REGION Network 268
   RUNG wire#powerrail
      Contact( "EMS".Carrier[02].SDC_OUT.HeartBeat )
      Coil( "Carrier_02_Heartbeat" )
   END_RUNG
   // the same network as SCL:
   "Carrier_02_Heartbeat" := "EMS".Carrier[02].SDC_OUT.HeartBeat;
END_REGION

REGION Network 269
   RUNG wire#powerrail
      Contact( "EMS".Carrier[02].SDC_OUT.DriveFwdCMD )
      I_Contact( "EMS".Carrier[01].SDC_IN.CrashDetectStatus )
      Coil( "Carrier_02_Drive_Forward_Command" )
   END_RUNG
   // the same network as SCL:
   "Carrier_02_Drive_Forward_Command" := "EMS".Carrier[02].SDC_OUT.DriveFwdCMD AND NOT "EMS".Carrier[01].SDC_IN.CrashDetectStatus;
END_REGION

REGION Network 270
   RUNG wire#powerrail
      Contact( "EMS".Carrier[02].SDC_OUT.FaultReset )
      Coil( "Carrier_02_Fault_Reset" )
   END_RUNG
   // the same network as SCL:
   "Carrier_02_Fault_Reset" := "EMS".Carrier[02].SDC_OUT.FaultReset;
END_REGION

REGION Network 271
   RUNG wire#powerrail
      Contact( "EMS".Carrier[02].SDC_OUT.AtCmdPos )
      Coil( "Carrier_02_At_Command_Position" )
   END_RUNG
   // the same network as SCL:
   "Carrier_02_At_Command_Position" := "EMS".Carrier[02].SDC_OUT.AtCmdPos;
END_REGION

REGION Network 272
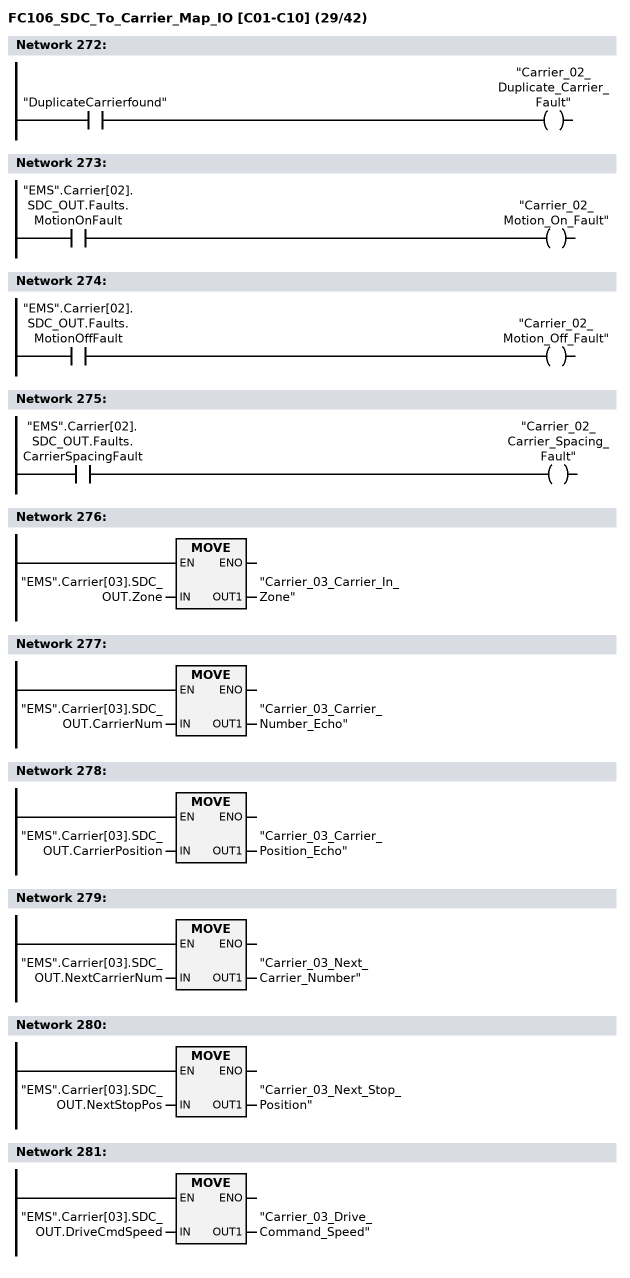
   RUNG wire#powerrail
      Contact( "DuplicateCarrierfound" )
      Coil( "Carrier_02_Duplicate_Carrier_Fault" )
   END_RUNG
   // the same network as SCL:
   "Carrier_02_Duplicate_Carrier_Fault" := "DuplicateCarrierfound";
END_REGION

REGION Network 273
   RUNG wire#powerrail
      Contact( "EMS".Carrier[02].SDC_OUT.Faults.MotionOnFault )
      Coil( "Carrier_02_Motion_On_Fault" )
   END_RUNG
   // the same network as SCL:
   "Carrier_02_Motion_On_Fault" := "EMS".Carrier[02].SDC_OUT.Faults.MotionOnFault;
END_REGION

REGION Network 274
   RUNG wire#powerrail
      Contact( "EMS".Carrier[02].SDC_OUT.Faults.MotionOffFault )
      Coil( "Carrier_02_Motion_Off_Fault" )
   END_RUNG
   // the same network as SCL:
   "Carrier_02_Motion_Off_Fault" := "EMS".Carrier[02].SDC_OUT.Faults.MotionOffFault;
END_REGION

REGION Network 275
   RUNG wire#powerrail
      Contact( "EMS".Carrier[02].SDC_OUT.Faults.CarrierSpacingFault )
      Coil( "Carrier_02_Carrier_Spacing_Fault" )
   END_RUNG
   // the same network as SCL:
   "Carrier_02_Carrier_Spacing_Fault" := "EMS".Carrier[02].SDC_OUT.Faults.CarrierSpacingFault;
END_REGION

REGION Network 276
   RUNG wire#powerrail
      Move(in := "EMS".Carrier[03].SDC_OUT.Zone, out1 => "Carrier_03_Carrier_In_Zone")
   END_RUNG
   // the same network as SCL:
   "Carrier_03_Carrier_In_Zone" := "EMS".Carrier[03].SDC_OUT.Zone;
END_REGION

REGION Network 277
   RUNG wire#powerrail
      Move(in := "EMS".Carrier[03].SDC_OUT.CarrierNum, out1 => "Carrier_03_Carrier_Number_Echo")
   END_RUNG
   // the same network as SCL:
   "Carrier_03_Carrier_Number_Echo" := "EMS".Carrier[03].SDC_OUT.CarrierNum;
END_REGION

REGION Network 278
   RUNG wire#powerrail
      Move(in := "EMS".Carrier[03].SDC_OUT.CarrierPosition, out1 => "Carrier_03_Carrier_Position_Echo")
   END_RUNG
   // the same network as SCL:
   "Carrier_03_Carrier_Position_Echo" := "EMS".Carrier[03].SDC_OUT.CarrierPosition;
END_REGION

REGION Network 279
   RUNG wire#powerrail
      Move(in := "EMS".Carrier[03].SDC_OUT.NextCarrierNum, out1 => "Carrier_03_Next_Carrier_Number")
   END_RUNG
   // the same network as SCL:
   "Carrier_03_Next_Carrier_Number" := "EMS".Carrier[03].SDC_OUT.NextCarrierNum;
END_REGION

REGION Network 280
   RUNG wire#powerrail
      Move(in := "EMS".Carrier[03].SDC_OUT.NextStopPos, out1 => "Carrier_03_Next_Stop_Position")
   END_RUNG
   // the same network as SCL:
   "Carrier_03_Next_Stop_Position" := "EMS".Carrier[03].SDC_OUT.NextStopPos;
END_REGION

REGION Network 281
   RUNG wire#powerrail
      Move(in := "EMS".Carrier[03].SDC_OUT.DriveCmdSpeed, out1 => "Carrier_03_Drive_Command_Speed")
   END_RUNG
   // the same network as SCL:
   "Carrier_03_Drive_Command_Speed" := "EMS".Carrier[03].SDC_OUT.DriveCmdSpeed;
END_REGION

REGION Network 282
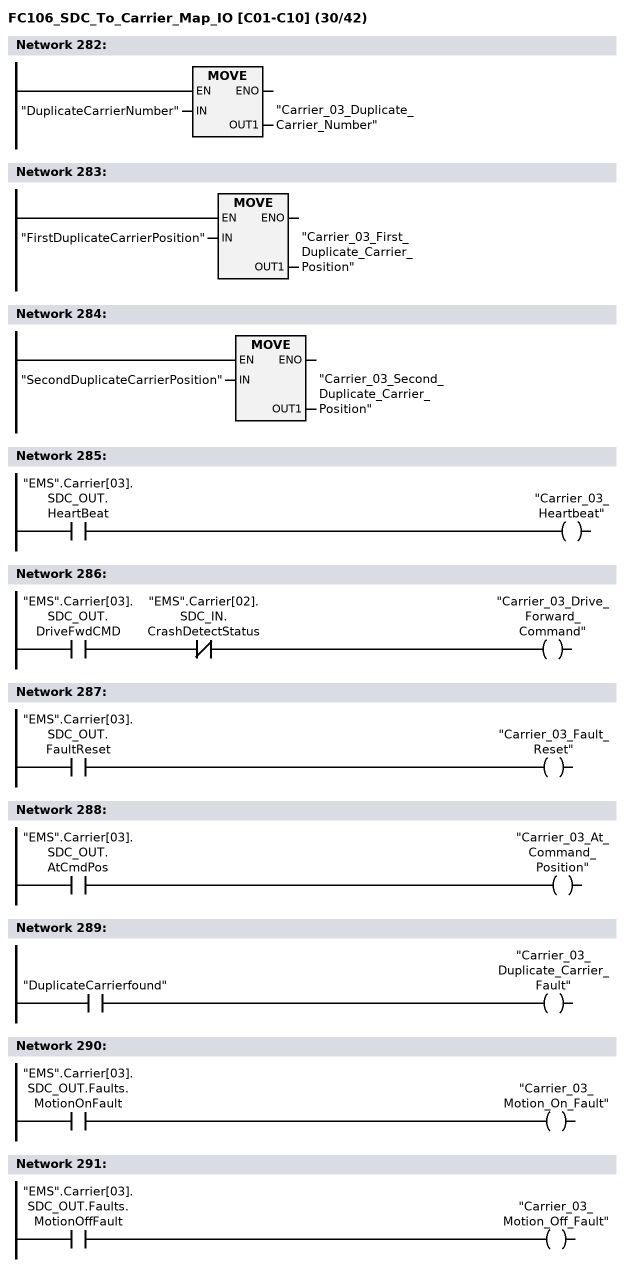
   RUNG wire#powerrail
      Move(in := "DuplicateCarrierNumber", out1 => "Carrier_03_Duplicate_Carrier_Number")
   END_RUNG
   // the same network as SCL:
   "Carrier_03_Duplicate_Carrier_Number" := "DuplicateCarrierNumber";
END_REGION

REGION Network 283
   RUNG wire#powerrail
      Move(in := "FirstDuplicateCarrierPosition", out1 => "Carrier_03_First_Duplicate_Carrier_Position")
   END_RUNG
   // the same network as SCL:
   "Carrier_03_First_Duplicate_Carrier_Position" := "FirstDuplicateCarrierPosition";
END_REGION

REGION Network 284
   RUNG wire#powerrail
      Move(in := "SecondDuplicateCarrierPosition", out1 => "Carrier_03_Second_Duplicate_Carrier_Position")
   END_RUNG
   // the same network as SCL:
   "Carrier_03_Second_Duplicate_Carrier_Position" := "SecondDuplicateCarrierPosition";
END_REGION

REGION Network 285
   RUNG wire#powerrail
      Contact( "EMS".Carrier[03].SDC_OUT.HeartBeat )
      Coil( "Carrier_03_Heartbeat" )
   END_RUNG
   // the same network as SCL:
   "Carrier_03_Heartbeat" := "EMS".Carrier[03].SDC_OUT.HeartBeat;
END_REGION

REGION Network 286
   RUNG wire#powerrail
      Contact( "EMS".Carrier[03].SDC_OUT.DriveFwdCMD )
      I_Contact( "EMS".Carrier[02].SDC_IN.CrashDetectStatus )
      Coil( "Carrier_03_Drive_Forward_Command" )
   END_RUNG
   // the same network as SCL:
   "Carrier_03_Drive_Forward_Command" := "EMS".Carrier[03].SDC_OUT.DriveFwdCMD AND NOT "EMS".Carrier[02].SDC_IN.CrashDetectStatus;
END_REGION

REGION Network 287
   RUNG wire#powerrail
      Contact( "EMS".Carrier[03].SDC_OUT.FaultReset )
      Coil( "Carrier_03_Fault_Reset" )
   END_RUNG
   // the same network as SCL:
   "Carrier_03_Fault_Reset" := "EMS".Carrier[03].SDC_OUT.FaultReset;
END_REGION

REGION Network 288
   RUNG wire#powerrail
      Contact( "EMS".Carrier[03].SDC_OUT.AtCmdPos )
      Coil( "Carrier_03_At_Command_Position" )
   END_RUNG
   // the same network as SCL:
   "Carrier_03_At_Command_Position" := "EMS".Carrier[03].SDC_OUT.AtCmdPos;
END_REGION

REGION Network 289
   RUNG wire#powerrail
      Contact( "DuplicateCarrierfound" )
      Coil( "Carrier_03_Duplicate_Carrier_Fault" )
   END_RUNG
   // the same network as SCL:
   "Carrier_03_Duplicate_Carrier_Fault" := "DuplicateCarrierfound";
END_REGION

REGION Network 290
   RUNG wire#powerrail
      Contact( "EMS".Carrier[03].SDC_OUT.Faults.MotionOnFault )
      Coil( "Carrier_03_Motion_On_Fault" )
   END_RUNG
   // the same network as SCL:
   "Carrier_03_Motion_On_Fault" := "EMS".Carrier[03].SDC_OUT.Faults.MotionOnFault;
END_REGION

REGION Network 291
   RUNG wire#powerrail
      Contact( "EMS".Carrier[03].SDC_OUT.Faults.MotionOffFault )
      Coil( "Carrier_03_Motion_Off_Fault" )
   END_RUNG
   // the same network as SCL:
   "Carrier_03_Motion_Off_Fault" := "EMS".Carrier[03].SDC_OUT.Faults.MotionOffFault;
END_REGION

REGION Network 292
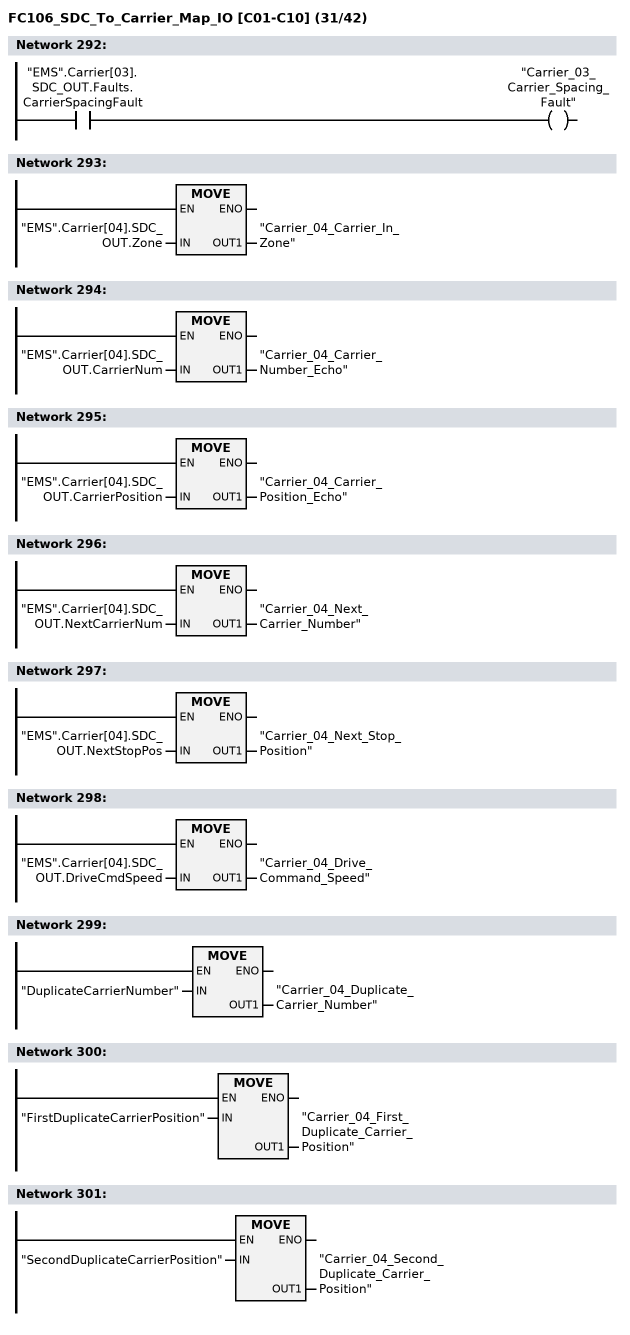
   RUNG wire#powerrail
      Contact( "EMS".Carrier[03].SDC_OUT.Faults.CarrierSpacingFault )
      Coil( "Carrier_03_Carrier_Spacing_Fault" )
   END_RUNG
   // the same network as SCL:
   "Carrier_03_Carrier_Spacing_Fault" := "EMS".Carrier[03].SDC_OUT.Faults.CarrierSpacingFault;
END_REGION

REGION Network 293
   RUNG wire#powerrail
      Move(in := "EMS".Carrier[04].SDC_OUT.Zone, out1 => "Carrier_04_Carrier_In_Zone")
   END_RUNG
   // the same network as SCL:
   "Carrier_04_Carrier_In_Zone" := "EMS".Carrier[04].SDC_OUT.Zone;
END_REGION

REGION Network 294
   RUNG wire#powerrail
      Move(in := "EMS".Carrier[04].SDC_OUT.CarrierNum, out1 => "Carrier_04_Carrier_Number_Echo")
   END_RUNG
   // the same network as SCL:
   "Carrier_04_Carrier_Number_Echo" := "EMS".Carrier[04].SDC_OUT.CarrierNum;
END_REGION

REGION Network 295
   RUNG wire#powerrail
      Move(in := "EMS".Carrier[04].SDC_OUT.CarrierPosition, out1 => "Carrier_04_Carrier_Position_Echo")
   END_RUNG
   // the same network as SCL:
   "Carrier_04_Carrier_Position_Echo" := "EMS".Carrier[04].SDC_OUT.CarrierPosition;
END_REGION

REGION Network 296
   RUNG wire#powerrail
      Move(in := "EMS".Carrier[04].SDC_OUT.NextCarrierNum, out1 => "Carrier_04_Next_Carrier_Number")
   END_RUNG
   // the same network as SCL:
   "Carrier_04_Next_Carrier_Number" := "EMS".Carrier[04].SDC_OUT.NextCarrierNum;
END_REGION

REGION Network 297
   RUNG wire#powerrail
      Move(in := "EMS".Carrier[04].SDC_OUT.NextStopPos, out1 => "Carrier_04_Next_Stop_Position")
   END_RUNG
   // the same network as SCL:
   "Carrier_04_Next_Stop_Position" := "EMS".Carrier[04].SDC_OUT.NextStopPos;
END_REGION

REGION Network 298
   RUNG wire#powerrail
      Move(in := "EMS".Carrier[04].SDC_OUT.DriveCmdSpeed, out1 => "Carrier_04_Drive_Command_Speed")
   END_RUNG
   // the same network as SCL:
   "Carrier_04_Drive_Command_Speed" := "EMS".Carrier[04].SDC_OUT.DriveCmdSpeed;
END_REGION

REGION Network 299
   RUNG wire#powerrail
      Move(in := "DuplicateCarrierNumber", out1 => "Carrier_04_Duplicate_Carrier_Number")
   END_RUNG
   // the same network as SCL:
   "Carrier_04_Duplicate_Carrier_Number" := "DuplicateCarrierNumber";
END_REGION

REGION Network 300
   RUNG wire#powerrail
      Move(in := "FirstDuplicateCarrierPosition", out1 => "Carrier_04_First_Duplicate_Carrier_Position")
   END_RUNG
   // the same network as SCL:
   "Carrier_04_First_Duplicate_Carrier_Position" := "FirstDuplicateCarrierPosition";
END_REGION

REGION Network 301
   RUNG wire#powerrail
      Move(in := "SecondDuplicateCarrierPosition", out1 => "Carrier_04_Second_Duplicate_Carrier_Position")
   END_RUNG
   // the same network as SCL:
   "Carrier_04_Second_Duplicate_Carrier_Position" := "SecondDuplicateCarrierPosition";
END_REGION

REGION Network 302
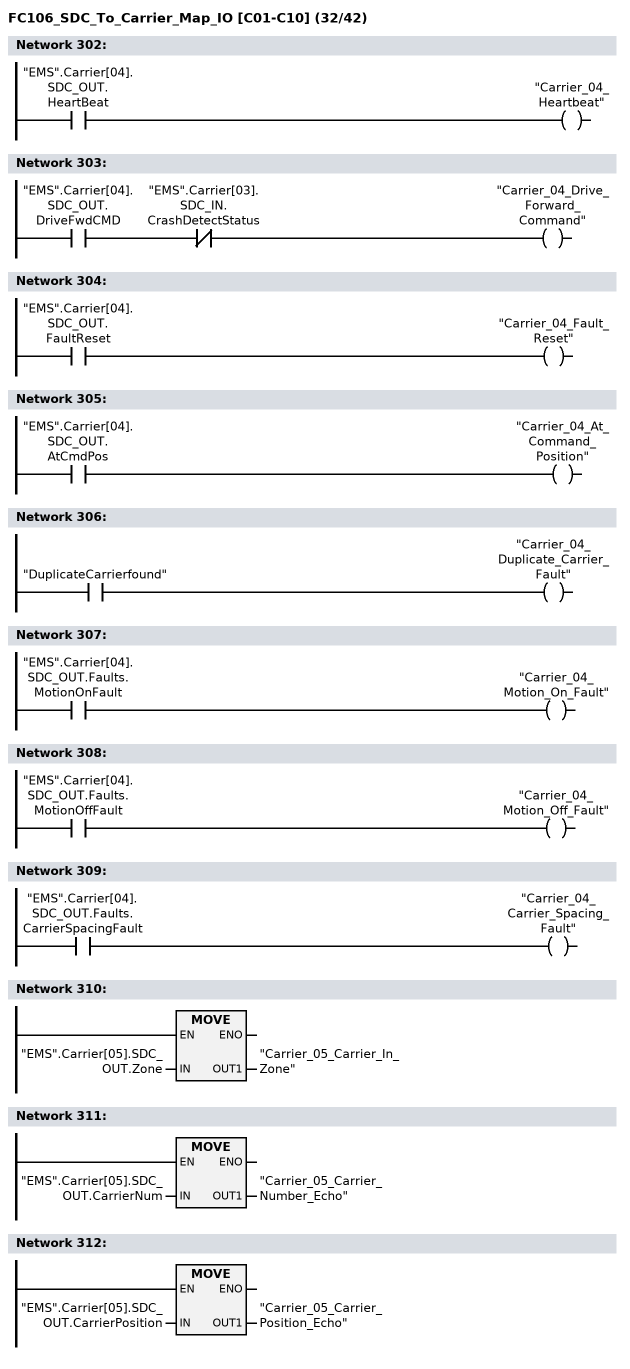
   RUNG wire#powerrail
      Contact( "EMS".Carrier[04].SDC_OUT.HeartBeat )
      Coil( "Carrier_04_Heartbeat" )
   END_RUNG
   // the same network as SCL:
   "Carrier_04_Heartbeat" := "EMS".Carrier[04].SDC_OUT.HeartBeat;
END_REGION

REGION Network 303
   RUNG wire#powerrail
      Contact( "EMS".Carrier[04].SDC_OUT.DriveFwdCMD )
      I_Contact( "EMS".Carrier[03].SDC_IN.CrashDetectStatus )
      Coil( "Carrier_04_Drive_Forward_Command" )
   END_RUNG
   // the same network as SCL:
   "Carrier_04_Drive_Forward_Command" := "EMS".Carrier[04].SDC_OUT.DriveFwdCMD AND NOT "EMS".Carrier[03].SDC_IN.CrashDetectStatus;
END_REGION

REGION Network 304
   RUNG wire#powerrail
      Contact( "EMS".Carrier[04].SDC_OUT.FaultReset )
      Coil( "Carrier_04_Fault_Reset" )
   END_RUNG
   // the same network as SCL:
   "Carrier_04_Fault_Reset" := "EMS".Carrier[04].SDC_OUT.FaultReset;
END_REGION

REGION Network 305
   RUNG wire#powerrail
      Contact( "EMS".Carrier[04].SDC_OUT.AtCmdPos )
      Coil( "Carrier_04_At_Command_Position" )
   END_RUNG
   // the same network as SCL:
   "Carrier_04_At_Command_Position" := "EMS".Carrier[04].SDC_OUT.AtCmdPos;
END_REGION

REGION Network 306
   RUNG wire#powerrail
      Contact( "DuplicateCarrierfound" )
      Coil( "Carrier_04_Duplicate_Carrier_Fault" )
   END_RUNG
   // the same network as SCL:
   "Carrier_04_Duplicate_Carrier_Fault" := "DuplicateCarrierfound";
END_REGION

REGION Network 307
   RUNG wire#powerrail
      Contact( "EMS".Carrier[04].SDC_OUT.Faults.MotionOnFault )
      Coil( "Carrier_04_Motion_On_Fault" )
   END_RUNG
   // the same network as SCL:
   "Carrier_04_Motion_On_Fault" := "EMS".Carrier[04].SDC_OUT.Faults.MotionOnFault;
END_REGION

REGION Network 308
   RUNG wire#powerrail
      Contact( "EMS".Carrier[04].SDC_OUT.Faults.MotionOffFault )
      Coil( "Carrier_04_Motion_Off_Fault" )
   END_RUNG
   // the same network as SCL:
   "Carrier_04_Motion_Off_Fault" := "EMS".Carrier[04].SDC_OUT.Faults.MotionOffFault;
END_REGION

REGION Network 309
   RUNG wire#powerrail
      Contact( "EMS".Carrier[04].SDC_OUT.Faults.CarrierSpacingFault )
      Coil( "Carrier_04_Carrier_Spacing_Fault" )
   END_RUNG
   // the same network as SCL:
   "Carrier_04_Carrier_Spacing_Fault" := "EMS".Carrier[04].SDC_OUT.Faults.CarrierSpacingFault;
END_REGION

REGION Network 310
   RUNG wire#powerrail
      Move(in := "EMS".Carrier[05].SDC_OUT.Zone, out1 => "Carrier_05_Carrier_In_Zone")
   END_RUNG
   // the same network as SCL:
   "Carrier_05_Carrier_In_Zone" := "EMS".Carrier[05].SDC_OUT.Zone;
END_REGION

REGION Network 311
   RUNG wire#powerrail
      Move(in := "EMS".Carrier[05].SDC_OUT.CarrierNum, out1 => "Carrier_05_Carrier_Number_Echo")
   END_RUNG
   // the same network as SCL:
   "Carrier_05_Carrier_Number_Echo" := "EMS".Carrier[05].SDC_OUT.CarrierNum;
END_REGION

REGION Network 312
   RUNG wire#powerrail
      Move(in := "EMS".Carrier[05].SDC_OUT.CarrierPosition, out1 => "Carrier_05_Carrier_Position_Echo")
   END_RUNG
   // the same network as SCL:
   "Carrier_05_Carrier_Position_Echo" := "EMS".Carrier[05].SDC_OUT.CarrierPosition;
END_REGION

REGION Network 313
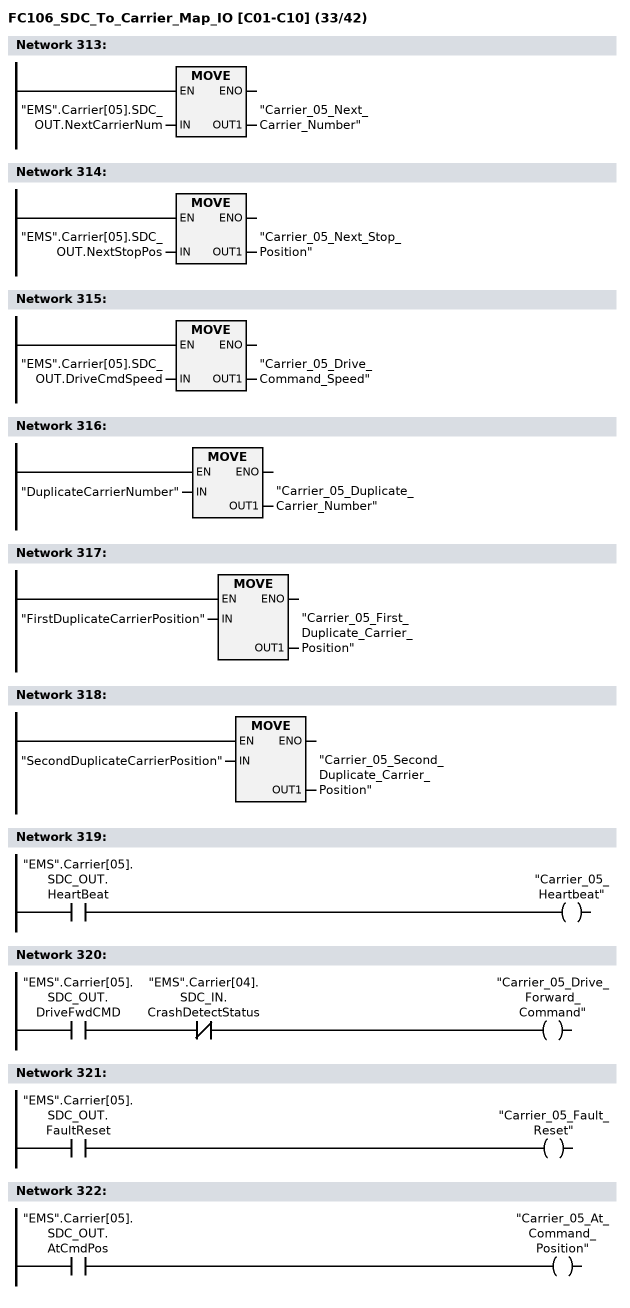
   RUNG wire#powerrail
      Move(in := "EMS".Carrier[05].SDC_OUT.NextCarrierNum, out1 => "Carrier_05_Next_Carrier_Number")
   END_RUNG
   // the same network as SCL:
   "Carrier_05_Next_Carrier_Number" := "EMS".Carrier[05].SDC_OUT.NextCarrierNum;
END_REGION

REGION Network 314
   RUNG wire#powerrail
      Move(in := "EMS".Carrier[05].SDC_OUT.NextStopPos, out1 => "Carrier_05_Next_Stop_Position")
   END_RUNG
   // the same network as SCL:
   "Carrier_05_Next_Stop_Position" := "EMS".Carrier[05].SDC_OUT.NextStopPos;
END_REGION

REGION Network 315
   RUNG wire#powerrail
      Move(in := "EMS".Carrier[05].SDC_OUT.DriveCmdSpeed, out1 => "Carrier_05_Drive_Command_Speed")
   END_RUNG
   // the same network as SCL:
   "Carrier_05_Drive_Command_Speed" := "EMS".Carrier[05].SDC_OUT.DriveCmdSpeed;
END_REGION

REGION Network 316
   RUNG wire#powerrail
      Move(in := "DuplicateCarrierNumber", out1 => "Carrier_05_Duplicate_Carrier_Number")
   END_RUNG
   // the same network as SCL:
   "Carrier_05_Duplicate_Carrier_Number" := "DuplicateCarrierNumber";
END_REGION

REGION Network 317
   RUNG wire#powerrail
      Move(in := "FirstDuplicateCarrierPosition", out1 => "Carrier_05_First_Duplicate_Carrier_Position")
   END_RUNG
   // the same network as SCL:
   "Carrier_05_First_Duplicate_Carrier_Position" := "FirstDuplicateCarrierPosition";
END_REGION

REGION Network 318
   RUNG wire#powerrail
      Move(in := "SecondDuplicateCarrierPosition", out1 => "Carrier_05_Second_Duplicate_Carrier_Position")
   END_RUNG
   // the same network as SCL:
   "Carrier_05_Second_Duplicate_Carrier_Position" := "SecondDuplicateCarrierPosition";
END_REGION

REGION Network 319
   RUNG wire#powerrail
      Contact( "EMS".Carrier[05].SDC_OUT.HeartBeat )
      Coil( "Carrier_05_Heartbeat" )
   END_RUNG
   // the same network as SCL:
   "Carrier_05_Heartbeat" := "EMS".Carrier[05].SDC_OUT.HeartBeat;
END_REGION

REGION Network 320
   RUNG wire#powerrail
      Contact( "EMS".Carrier[05].SDC_OUT.DriveFwdCMD )
      I_Contact( "EMS".Carrier[04].SDC_IN.CrashDetectStatus )
      Coil( "Carrier_05_Drive_Forward_Command" )
   END_RUNG
   // the same network as SCL:
   "Carrier_05_Drive_Forward_Command" := "EMS".Carrier[05].SDC_OUT.DriveFwdCMD AND NOT "EMS".Carrier[04].SDC_IN.CrashDetectStatus;
END_REGION

REGION Network 321
   RUNG wire#powerrail
      Contact( "EMS".Carrier[05].SDC_OUT.FaultReset )
      Coil( "Carrier_05_Fault_Reset" )
   END_RUNG
   // the same network as SCL:
   "Carrier_05_Fault_Reset" := "EMS".Carrier[05].SDC_OUT.FaultReset;
END_REGION

REGION Network 322
   RUNG wire#powerrail
      Contact( "EMS".Carrier[05].SDC_OUT.AtCmdPos )
      Coil( "Carrier_05_At_Command_Position" )
   END_RUNG
   // the same network as SCL:
   "Carrier_05_At_Command_Position" := "EMS".Carrier[05].SDC_OUT.AtCmdPos;
END_REGION

REGION Network 323
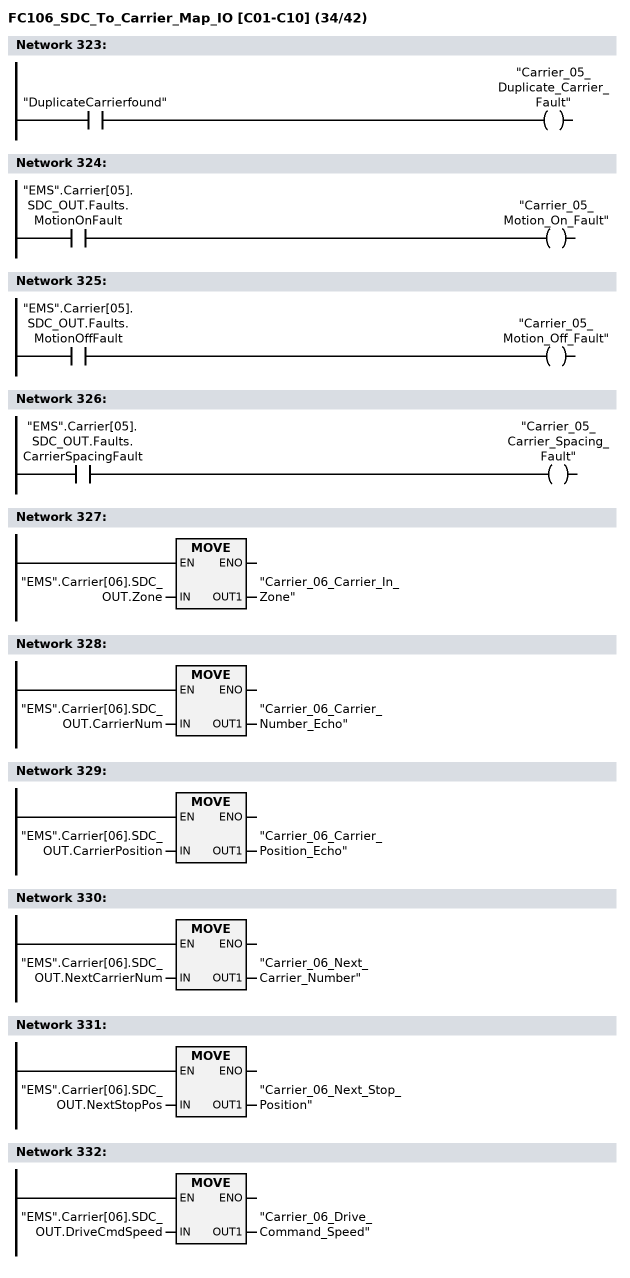
   RUNG wire#powerrail
      Contact( "DuplicateCarrierfound" )
      Coil( "Carrier_05_Duplicate_Carrier_Fault" )
   END_RUNG
   // the same network as SCL:
   "Carrier_05_Duplicate_Carrier_Fault" := "DuplicateCarrierfound";
END_REGION

REGION Network 324
   RUNG wire#powerrail
      Contact( "EMS".Carrier[05].SDC_OUT.Faults.MotionOnFault )
      Coil( "Carrier_05_Motion_On_Fault" )
   END_RUNG
   // the same network as SCL:
   "Carrier_05_Motion_On_Fault" := "EMS".Carrier[05].SDC_OUT.Faults.MotionOnFault;
END_REGION

REGION Network 325
   RUNG wire#powerrail
      Contact( "EMS".Carrier[05].SDC_OUT.Faults.MotionOffFault )
      Coil( "Carrier_05_Motion_Off_Fault" )
   END_RUNG
   // the same network as SCL:
   "Carrier_05_Motion_Off_Fault" := "EMS".Carrier[05].SDC_OUT.Faults.MotionOffFault;
END_REGION

REGION Network 326
   RUNG wire#powerrail
      Contact( "EMS".Carrier[05].SDC_OUT.Faults.CarrierSpacingFault )
      Coil( "Carrier_05_Carrier_Spacing_Fault" )
   END_RUNG
   // the same network as SCL:
   "Carrier_05_Carrier_Spacing_Fault" := "EMS".Carrier[05].SDC_OUT.Faults.CarrierSpacingFault;
END_REGION

REGION Network 327
   RUNG wire#powerrail
      Move(in := "EMS".Carrier[06].SDC_OUT.Zone, out1 => "Carrier_06_Carrier_In_Zone")
   END_RUNG
   // the same network as SCL:
   "Carrier_06_Carrier_In_Zone" := "EMS".Carrier[06].SDC_OUT.Zone;
END_REGION

REGION Network 328
   RUNG wire#powerrail
      Move(in := "EMS".Carrier[06].SDC_OUT.CarrierNum, out1 => "Carrier_06_Carrier_Number_Echo")
   END_RUNG
   // the same network as SCL:
   "Carrier_06_Carrier_Number_Echo" := "EMS".Carrier[06].SDC_OUT.CarrierNum;
END_REGION

REGION Network 329
   RUNG wire#powerrail
      Move(in := "EMS".Carrier[06].SDC_OUT.CarrierPosition, out1 => "Carrier_06_Carrier_Position_Echo")
   END_RUNG
   // the same network as SCL:
   "Carrier_06_Carrier_Position_Echo" := "EMS".Carrier[06].SDC_OUT.CarrierPosition;
END_REGION

REGION Network 330
   RUNG wire#powerrail
      Move(in := "EMS".Carrier[06].SDC_OUT.NextCarrierNum, out1 => "Carrier_06_Next_Carrier_Number")
   END_RUNG
   // the same network as SCL:
   "Carrier_06_Next_Carrier_Number" := "EMS".Carrier[06].SDC_OUT.NextCarrierNum;
END_REGION

REGION Network 331
   RUNG wire#powerrail
      Move(in := "EMS".Carrier[06].SDC_OUT.NextStopPos, out1 => "Carrier_06_Next_Stop_Position")
   END_RUNG
   // the same network as SCL:
   "Carrier_06_Next_Stop_Position" := "EMS".Carrier[06].SDC_OUT.NextStopPos;
END_REGION

REGION Network 332
   RUNG wire#powerrail
      Move(in := "EMS".Carrier[06].SDC_OUT.DriveCmdSpeed, out1 => "Carrier_06_Drive_Command_Speed")
   END_RUNG
   // the same network as SCL:
   "Carrier_06_Drive_Command_Speed" := "EMS".Carrier[06].SDC_OUT.DriveCmdSpeed;
END_REGION

REGION Network 333
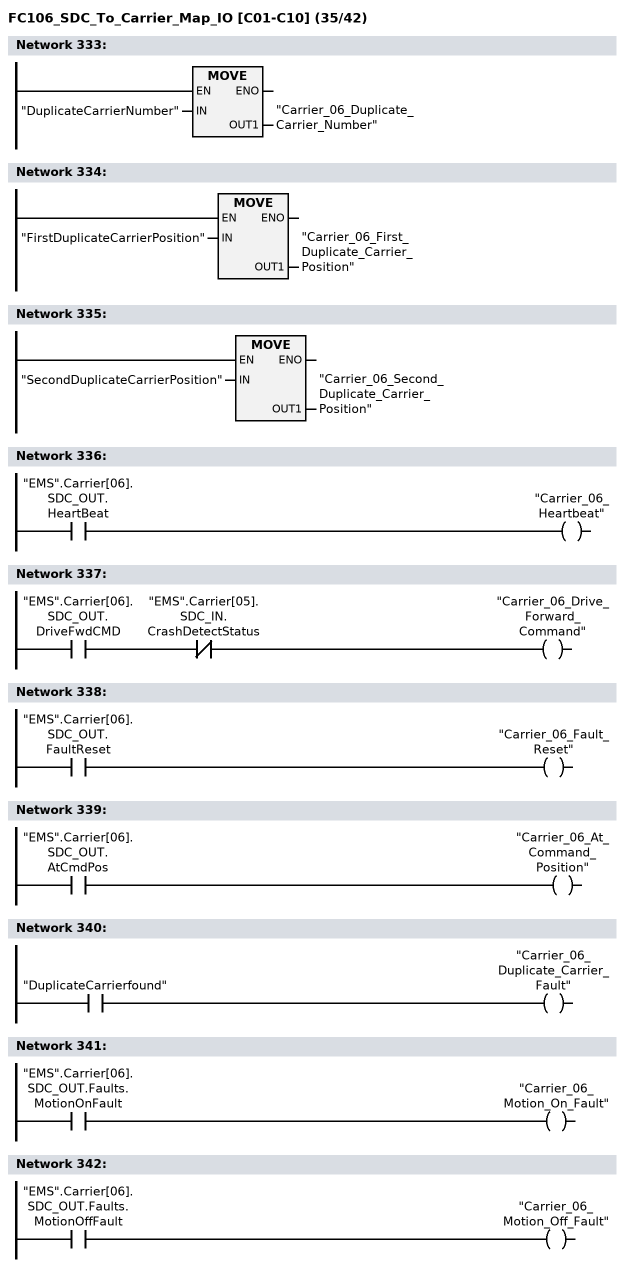
   RUNG wire#powerrail
      Move(in := "DuplicateCarrierNumber", out1 => "Carrier_06_Duplicate_Carrier_Number")
   END_RUNG
   // the same network as SCL:
   "Carrier_06_Duplicate_Carrier_Number" := "DuplicateCarrierNumber";
END_REGION

REGION Network 334
   RUNG wire#powerrail
      Move(in := "FirstDuplicateCarrierPosition", out1 => "Carrier_06_First_Duplicate_Carrier_Position")
   END_RUNG
   // the same network as SCL:
   "Carrier_06_First_Duplicate_Carrier_Position" := "FirstDuplicateCarrierPosition";
END_REGION

REGION Network 335
   RUNG wire#powerrail
      Move(in := "SecondDuplicateCarrierPosition", out1 => "Carrier_06_Second_Duplicate_Carrier_Position")
   END_RUNG
   // the same network as SCL:
   "Carrier_06_Second_Duplicate_Carrier_Position" := "SecondDuplicateCarrierPosition";
END_REGION

REGION Network 336
   RUNG wire#powerrail
      Contact( "EMS".Carrier[06].SDC_OUT.HeartBeat )
      Coil( "Carrier_06_Heartbeat" )
   END_RUNG
   // the same network as SCL:
   "Carrier_06_Heartbeat" := "EMS".Carrier[06].SDC_OUT.HeartBeat;
END_REGION

REGION Network 337
   RUNG wire#powerrail
      Contact( "EMS".Carrier[06].SDC_OUT.DriveFwdCMD )
      I_Contact( "EMS".Carrier[05].SDC_IN.CrashDetectStatus )
      Coil( "Carrier_06_Drive_Forward_Command" )
   END_RUNG
   // the same network as SCL:
   "Carrier_06_Drive_Forward_Command" := "EMS".Carrier[06].SDC_OUT.DriveFwdCMD AND NOT "EMS".Carrier[05].SDC_IN.CrashDetectStatus;
END_REGION

REGION Network 338
   RUNG wire#powerrail
      Contact( "EMS".Carrier[06].SDC_OUT.FaultReset )
      Coil( "Carrier_06_Fault_Reset" )
   END_RUNG
   // the same network as SCL:
   "Carrier_06_Fault_Reset" := "EMS".Carrier[06].SDC_OUT.FaultReset;
END_REGION

REGION Network 339
   RUNG wire#powerrail
      Contact( "EMS".Carrier[06].SDC_OUT.AtCmdPos )
      Coil( "Carrier_06_At_Command_Position" )
   END_RUNG
   // the same network as SCL:
   "Carrier_06_At_Command_Position" := "EMS".Carrier[06].SDC_OUT.AtCmdPos;
END_REGION

REGION Network 340
   RUNG wire#powerrail
      Contact( "DuplicateCarrierfound" )
      Coil( "Carrier_06_Duplicate_Carrier_Fault" )
   END_RUNG
   // the same network as SCL:
   "Carrier_06_Duplicate_Carrier_Fault" := "DuplicateCarrierfound";
END_REGION

REGION Network 341
   RUNG wire#powerrail
      Contact( "EMS".Carrier[06].SDC_OUT.Faults.MotionOnFault )
      Coil( "Carrier_06_Motion_On_Fault" )
   END_RUNG
   // the same network as SCL:
   "Carrier_06_Motion_On_Fault" := "EMS".Carrier[06].SDC_OUT.Faults.MotionOnFault;
END_REGION

REGION Network 342
   RUNG wire#powerrail
      Contact( "EMS".Carrier[06].SDC_OUT.Faults.MotionOffFault )
      Coil( "Carrier_06_Motion_Off_Fault" )
   END_RUNG
   // the same network as SCL:
   "Carrier_06_Motion_Off_Fault" := "EMS".Carrier[06].SDC_OUT.Faults.MotionOffFault;
END_REGION

REGION Network 343
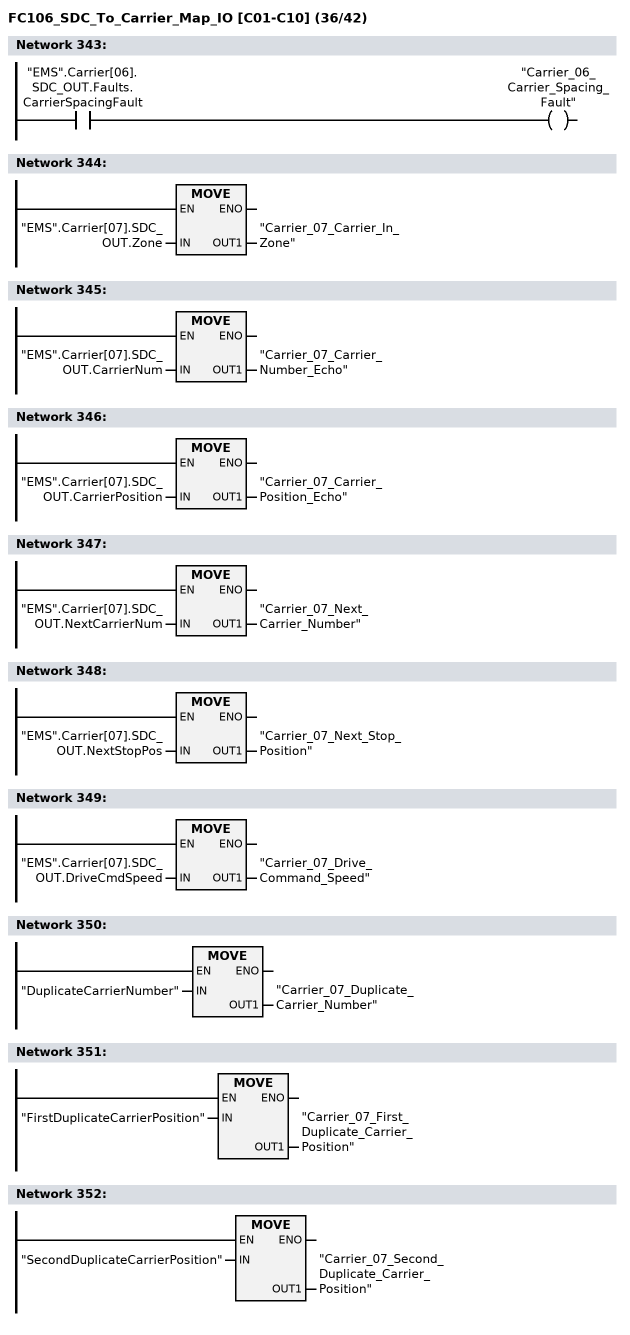
   RUNG wire#powerrail
      Contact( "EMS".Carrier[06].SDC_OUT.Faults.CarrierSpacingFault )
      Coil( "Carrier_06_Carrier_Spacing_Fault" )
   END_RUNG
   // the same network as SCL:
   "Carrier_06_Carrier_Spacing_Fault" := "EMS".Carrier[06].SDC_OUT.Faults.CarrierSpacingFault;
END_REGION

REGION Network 344
   RUNG wire#powerrail
      Move(in := "EMS".Carrier[07].SDC_OUT.Zone, out1 => "Carrier_07_Carrier_In_Zone")
   END_RUNG
   // the same network as SCL:
   "Carrier_07_Carrier_In_Zone" := "EMS".Carrier[07].SDC_OUT.Zone;
END_REGION

REGION Network 345
   RUNG wire#powerrail
      Move(in := "EMS".Carrier[07].SDC_OUT.CarrierNum, out1 => "Carrier_07_Carrier_Number_Echo")
   END_RUNG
   // the same network as SCL:
   "Carrier_07_Carrier_Number_Echo" := "EMS".Carrier[07].SDC_OUT.CarrierNum;
END_REGION

REGION Network 346
   RUNG wire#powerrail
      Move(in := "EMS".Carrier[07].SDC_OUT.CarrierPosition, out1 => "Carrier_07_Carrier_Position_Echo")
   END_RUNG
   // the same network as SCL:
   "Carrier_07_Carrier_Position_Echo" := "EMS".Carrier[07].SDC_OUT.CarrierPosition;
END_REGION

REGION Network 347
   RUNG wire#powerrail
      Move(in := "EMS".Carrier[07].SDC_OUT.NextCarrierNum, out1 => "Carrier_07_Next_Carrier_Number")
   END_RUNG
   // the same network as SCL:
   "Carrier_07_Next_Carrier_Number" := "EMS".Carrier[07].SDC_OUT.NextCarrierNum;
END_REGION

REGION Network 348
   RUNG wire#powerrail
      Move(in := "EMS".Carrier[07].SDC_OUT.NextStopPos, out1 => "Carrier_07_Next_Stop_Position")
   END_RUNG
   // the same network as SCL:
   "Carrier_07_Next_Stop_Position" := "EMS".Carrier[07].SDC_OUT.NextStopPos;
END_REGION

REGION Network 349
   RUNG wire#powerrail
      Move(in := "EMS".Carrier[07].SDC_OUT.DriveCmdSpeed, out1 => "Carrier_07_Drive_Command_Speed")
   END_RUNG
   // the same network as SCL:
   "Carrier_07_Drive_Command_Speed" := "EMS".Carrier[07].SDC_OUT.DriveCmdSpeed;
END_REGION

REGION Network 350
   RUNG wire#powerrail
      Move(in := "DuplicateCarrierNumber", out1 => "Carrier_07_Duplicate_Carrier_Number")
   END_RUNG
   // the same network as SCL:
   "Carrier_07_Duplicate_Carrier_Number" := "DuplicateCarrierNumber";
END_REGION

REGION Network 351
   RUNG wire#powerrail
      Move(in := "FirstDuplicateCarrierPosition", out1 => "Carrier_07_First_Duplicate_Carrier_Position")
   END_RUNG
   // the same network as SCL:
   "Carrier_07_First_Duplicate_Carrier_Position" := "FirstDuplicateCarrierPosition";
END_REGION

REGION Network 352
   RUNG wire#powerrail
      Move(in := "SecondDuplicateCarrierPosition", out1 => "Carrier_07_Second_Duplicate_Carrier_Position")
   END_RUNG
   // the same network as SCL:
   "Carrier_07_Second_Duplicate_Carrier_Position" := "SecondDuplicateCarrierPosition";
END_REGION

REGION Network 353